ScreenModuleEditorView "IO Field: Single Width; Stacked" 178x111
   IOField "tfLable" at 0,55 size 178x56; FormatPattern ????????????????????????????????????????
      on OnFinishInput: SetBit("Interface.inputFinished")
      Appearance <- "Interface.animate"
      Visibility <- "Interface.visible"
      ProcessValue <- "Interface.value"
      ObjectEnable <- "Interface.enable"
   TextField "iofData" at 0,0 size 178x55; Text 'Text'
      Visibility <- "Interface.visible"
*)

(* ===== HMI "HMI_RT_1" =====
system functions are stored by id; their names below are inferred from use

ScreenModuleEditorView "IO Field: Double Width; Stacked" 370x111
   IOField "tfLable" at 0,55 size 370x56; FormatPattern ????????????????????????????????????????
      on OnFinishInput: SetBit("Interface.inputFinished")
      Appearance <- "Interface.animate"
      ProcessValue <- "Interface.value"
      Visibility <- "Interface.visible"
      ObjectEnable <- "Interface.enable"
   TextField "iofData" at 0,0 size 370x55; Text 'Text'
      Visibility <- "Interface.visible"
*)

(* ===== HMI "HMI_RT_1" =====
system functions are stored by id; their names below are inferred from use

ScreenModuleEditorView "PB: Graphic/Text List" 65x45
   Button "Previous Station Group" at 0,0 size 65x45; TextOff 'Text'
      on Press: function_b14e0dd5("Interface.actuate", 0)
      Visibility <- "Interface.animate"
      ObjectEnable <- "Interface.animate"
      Appearance <- "Interface.animate"
*)

(* ===== HMI "HMI_RT_1" =====
system functions are stored by id; their names below are inferred from use

ScreenModuleEditorView "PB: Graphic/Text List" 65x45
   Button "Previous Station Group" at 0,0 size 65x45; TextOff 'Text'
      on Press: function_b14e0dd5("Interface.actuate", 0)
      Visibility <- "Interface.animate"
      ObjectEnable <- "Interface.animate"
      Appearance <- "Interface.animate"
*)

(* ===== HMI "HMI_RT_1" =====
system functions are stored by id; their names below are inferred from use

ScreenModuleEditorView "PB: Station Comm Status (Text Label)" 180x25
   Button "Station Select" at 0,0 size 180x25; TextOff 'Text'
      on Press: function_b14e0dd5("Interface.actuate", 0)
      Appearance <- "Interface.animate"
      ObjectEnable <- "Interface.enable"
      Visibility <- "Interface.visible"
*)

(* ===== HMI "HMI_RT_1" =====
system functions are stored by id; their names below are inferred from use

ScreenModuleEditorView "PB: Graphic/Text List" 65x45
   Button "Previous Station Group" at 0,0 size 65x45; TextOff 'Text'
      on Press: function_b14e0dd5("Interface.actuate", 0)
      Visibility <- "Interface.animate"
      ObjectEnable <- "Interface.animate"
      Appearance <- "Interface.animate"
*)

(* ===== HMI "HMI_RT_1" =====
system functions are stored by id; their names below are inferred from use

graphic list "Top": 0 '100 x 100 Top'; 1 '100 x 100 Actuated Top'

graphic list "Page Up": 0 '100 x 100 Page Up'; 1 '100 x 100 Actuated Page Up'

graphic list "Line Up": 0 '100 x 100 Line Up'; 1 '100 x 100 Actuated Line Up'

graphic list "Line Down": 0 '100 x 100 Line Down'; 1 '100 x 100 Actuated Line Down'

graphic list "Page Down": 0 '100 x 100 Page Down'; 1 '100 x 100 Actuated Page Down'

graphic list "Bottom": 0 '100 x 100 Bottom'; 1 '100 x 100 Actuated Bottom'

ScreenModuleEditorView "Nav Bar: Horizontal" 600x100
   Button "btnTop" at 1,1 size 98x98; TextOff 'Text'; PictureList "Top"
      on Press: function_b14e0dd5("Interface.top.actuate", 0)
      Visibility <- "Interface.top.visible"
      ObjectEnable <- "Interface.top.enable"
      ProcessValue <- "Interface.top.listSelect"
      Appearance <- "Interface.top.animate"
   Button "btnPageUp" at 101,1 size 98x98; TextOff 'Text'; PictureList "Page Up"
      on Press: function_b14e0dd5("Interface.pageUp.actuate", 0)
      Appearance <- "Interface.pageUp.animate"
      ObjectEnable <- "Interface.pageUp.enable"
      ProcessValue <- "Interface.pageUp.listSelect"
      Visibility <- "Interface.pageUp.visible"
   Button "btnLineUp" at 201,1 size 98x98; TextOff 'Text'; PictureList "Line Up"
      on Press: function_b14e0dd5("Interface.lineUp.actuate", 0)
      Visibility <- "Interface.lineUp.visible"
      ObjectEnable <- "Interface.lineUp.enable"
      ProcessValue <- "Interface.lineUp.listSelect"
      Appearance <- "Interface.lineUp.animate"
   Button "btnLineDown" at 301,1 size 98x98; TextOff 'Text'; PictureList "Line Down"
      on Press: function_b14e0dd5("Interface.lineUp.actuate", 0)
      Appearance <- "Interface.lineDown.animate"
      ObjectEnable <- "Interface.lineDown.enable"
      ProcessValue <- "Interface.lineDown.listSelect"
      Visibility <- "Interface.lineDown.visible"
   Button "btnPageDown" at 401,1 size 98x98; TextOff 'Text'; PictureList "Page Down"
      on Press: function_b14e0dd5("Interface.pageDown.actuate", 0)
      Visibility <- "Interface.pageDown.visible"
      ObjectEnable <- "Interface.pageDown.enable"
      ProcessValue <- "Interface.pageDown.listSelect"
      Appearance <- "Interface.pageDown.animate"
   Button "btnBottom" at 501,1 size 98x98; TextOff 'Text'; PictureList "Bottom"
      on Press: function_b14e0dd5("Interface.pageDown.actuate", 0)
      Appearance <- "Interface.bottom.animate"
      ObjectEnable <- "Interface.bottom.enable"
      ProcessValue <- "Interface.bottom.listSelect"
      Visibility <- "Interface.bottom.visible"
*)

(* ===== HMI "HMI_RT_1" =====
system functions are stored by id; their names below are inferred from use

graphic list "Top": 0 '100 x 100 Top'; 1 '100 x 100 Actuated Top'

graphic list "Page Up": 0 '100 x 100 Page Up'; 1 '100 x 100 Actuated Page Up'

graphic list "Line Up": 0 '100 x 100 Line Up'; 1 '100 x 100 Actuated Line Up'

graphic list "Line Down": 0 '100 x 100 Line Down'; 1 '100 x 100 Actuated Line Down'

graphic list "Page Down": 0 '100 x 100 Page Down'; 1 '100 x 100 Actuated Page Down'

graphic list "Bottom": 0 '100 x 100 Bottom'; 1 '100 x 100 Actuated Bottom'

ScreenModuleEditorView "Nav Bar: Horizontal" 600x100
   Button "btnTop" at 1,1 size 98x98; TextOff 'Text'; PictureList "Top"
      on Press: function_b14e0dd5("Interface.top_actuate", 0)
      Appearance <- "Interface.top_animate"
      ObjectEnable <- "Interface.top_enable"
      Visibility <- "Interface.top_visible"
   Button "btnPageUp" at 101,1 size 98x98; TextOff 'Text'; PictureList "Page Up"
      on Press: function_b14e0dd5("Interface.page_up_actuate", 0)
      Visibility <- "Interface.page_up_visible"
      ObjectEnable <- "Interface.page_up_enable"
      Appearance <- "Interface.page_up_animate"
   Button "btnLineUp" at 201,1 size 98x98; TextOff 'Text'; PictureList "Line Up"
      on Press: function_b14e0dd5("Interface.line_up_actuate", 0)
      Visibility <- "Interface.line_up_visible"
      ObjectEnable <- "Interface.line_up_enable"
      Appearance <- "Interface.line_up_animate"
   Button "btnLineDown" at 301,1 size 98x98; TextOff 'Text'; PictureList "Line Down"
      on Press: function_b14e0dd5("Interface.line_down_actuate", 0)
      Appearance <- "Interface.line_down_animate"
      ObjectEnable <- "Interface.line_down_enable"
      Visibility <- "Interface.line_down_visible"
   Button "btnPageDown" at 401,1 size 98x98; TextOff 'Text'; PictureList "Page Down"
      on Press: function_b14e0dd5("Interface.page_down_actuate", 0)
      Visibility <- "Interface.page_down_visible"
      ObjectEnable <- "Interface.page_down_enable"
      Appearance <- "Interface.page_down_animate"
   Button "btnBottom" at 501,1 size 98x98; TextOff 'Text'; PictureList "Bottom"
      on Press: function_b14e0dd5("Interface.botttom_actuate", 0)
      Appearance <- "Interface.botttom_animate"
      ObjectEnable <- "Interface.botttom_enable"
      Visibility <- "Interface.botttom_visible"
*)

(* ===== HMI "HMI_RT_1" =====
system functions are stored by id; their names below are inferred from use

graphic list "Top": 0 '100 x 100 Top'; 1 '100 x 100 Actuated Top'

graphic list "Page Up": 0 '100 x 100 Page Up'; 1 '100 x 100 Actuated Page Up'

graphic list "Line Up": 0 '100 x 100 Line Up'; 1 '100 x 100 Actuated Line Up'

graphic list "Line Down": 0 '100 x 100 Line Down'; 1 '100 x 100 Actuated Line Down'

graphic list "Page Down": 0 '100 x 100 Page Down'; 1 '100 x 100 Actuated Page Down'

graphic list "Bottom": 0 '100 x 100 Bottom'; 1 '100 x 100 Actuated Bottom'

ScreenModuleEditorView "Nav Bar: Vertical" 100x600
   Button "btnTop" at 1,1 size 98x98; TextOff 'Text'; PictureList "Top"
      on Press: function_b14e0dd5("Interface.top_actuate", 0)
      Appearance <- "Interface.top_animate"
      ObjectEnable <- "Interface.top_enable"
      Visibility <- "Interface.top_visible"
   Button "btnPageUp" at 1,101 size 98x98; TextOff 'Text'; PictureList "Page Up"
      on Press: function_b14e0dd5("Interface.page_up_actuate", 0)
      Visibility <- "Interface.page_up_visible"
      ObjectEnable <- "Interface.page_up_enable"
      Appearance <- "Interface.page_up_animate"
   Button "btnLineUp" at 1,201 size 98x98; TextOff 'Text'; PictureList "Line Up"
      on Press: function_b14e0dd5("Interface.line_up_actuate", 0)
      Appearance <- "Interface.line_up_animate"
      ObjectEnable <- "Interface.line_up_enable"
      Visibility <- "Interface.line_up_visible"
   Button "btnLineDown" at 1,301 size 98x98; TextOff 'Text'; PictureList "Line Down"
      on Press: function_b14e0dd5("Interface.line_down_actuate", 0)
      Visibility <- "Interface.line_down_visible"
      ObjectEnable <- "Interface.line_down_enable"
      Appearance <- "Interface.line_down_animate"
   Button "btnPageDown" at 1,401 size 98x98; TextOff 'Text'; PictureList "Page Down"
      on Press: function_b14e0dd5("Interface.page_down_actuate", 0)
      Appearance <- "Interface.page_down_animate"
      ObjectEnable <- "Interface.page_down_enable"
      Visibility <- "Interface.page_down_visible"
   Button "btnBottom" at 1,501 size 98x98; TextOff 'Text'; PictureList "Bottom"
      on Press: SetBit("Interface.bottom_actuate")
      Visibility <- "Interface.bottom_visible"
      ObjectEnable <- "Interface.bottom_enable"
      Appearance <- "Interface.bottom_animate"
*)

(* ===== HMI "HMI_RT_1" =====
system functions are stored by id; their names below are inferred from use

graphic list "Top": 0 '100 x 100 Top'; 1 '100 x 100 Actuated Top'

graphic list "Page Up": 0 '100 x 100 Page Up'; 1 '100 x 100 Actuated Page Up'

graphic list "Line Up": 0 '100 x 100 Line Up'; 1 '100 x 100 Actuated Line Up'

graphic list "Line Down": 0 '100 x 100 Line Down'; 1 '100 x 100 Actuated Line Down'

graphic list "Page Down": 0 '100 x 100 Page Down'; 1 '100 x 100 Actuated Page Down'

graphic list "Bottom": 0 '100 x 100 Bottom'; 1 '100 x 100 Actuated Bottom'

ScreenModuleEditorView "Nav Bar: Horizontal" 600x100
   Button "btnTop" at 1,1 size 98x98; TextOff 'Text'; PictureList "Top"
      on Press: function_b14e0dd5("Interface.top_actuate", 0)
      Appearance <- "Interface.top_animate"
      ObjectEnable <- "Interface.top_enable"
      Visibility <- "Interface.top_visible"
   Button "btnPageUp" at 101,1 size 98x98; TextOff 'Text'; PictureList "Page Up"
      on Press: function_b14e0dd5("Interface.page_up_actuate", 0)
      Visibility <- "Interface.page_up_visible"
      ObjectEnable <- "Interface.page_up_enable"
      Appearance <- "Interface.page_up_animate"
   Button "btnLineUp" at 201,1 size 98x98; TextOff 'Text'; PictureList "Line Up"
      on Press: function_b14e0dd5("Interface.line_up_actuate", 0)
      Visibility <- "Interface.line_up_visible"
      ObjectEnable <- "Interface.line_up_enable"
      Appearance <- "Interface.line_up_animate"
   Button "btnLineDown" at 301,1 size 98x98; TextOff 'Text'; PictureList "Line Down"
      on Press: function_b14e0dd5("Interface.line_down_actuate", 0)
      Appearance <- "Interface.line_down_animate"
      ObjectEnable <- "Interface.line_down_enable"
      Visibility <- "Interface.line_down_visible"
   Button "btnPageDown" at 401,1 size 98x98; TextOff 'Text'; PictureList "Page Down"
      on Press: function_b14e0dd5("Interface.page_down_actuate", 0)
      Visibility <- "Interface.page_down_visible"
      ObjectEnable <- "Interface.page_down_enable"
      Appearance <- "Interface.page_down_animate"
   Button "btnBottom" at 501,1 size 98x98; TextOff 'Text'; PictureList "Bottom"
      on Press: function_b14e0dd5("Interface.bottom_actuate", 0)
      Visibility <- "Interface.bottom_visible"
      ObjectEnable <- "Interface.bottom_enable"
      Appearance <- "Interface.bottom_animate"
*)

(* ===== HMI "HMI_RT_1" =====
system functions are stored by id; their names below are inferred from use

graphic list "Top": 0 '100 x 100 Top'; 1 '100 x 100 Actuated Top'

graphic list "Page Up": 0 '100 x 100 Page Up'; 1 '100 x 100 Actuated Page Up'

graphic list "Line Up": 0 '100 x 100 Line Up'; 1 '100 x 100 Actuated Line Up'

graphic list "Line Down": 0 '100 x 100 Line Down'; 1 '100 x 100 Actuated Line Down'

graphic list "Page Down": 0 '100 x 100 Page Down'; 1 '100 x 100 Actuated Page Down'

graphic list "Bottom": 0 '100 x 100 Bottom'; 1 '100 x 100 Actuated Bottom'

ScreenModuleEditorView "Nav Bar: Horizontal" 600x100
   Button "btnTop" at 1,1 size 98x98; TextOff 'Text'; PictureList "Top"
      on Press: function_b14e0dd5("Interface.top_actuate", 0)
      Appearance <- "Interface.top_animate"
      ObjectEnable <- "Interface.top_enable"
      Visibility <- "Interface.top_visible"
      ProcessValue <- "Interface.top_list_select"
   Button "btnPageUp" at 101,1 size 98x98; TextOff 'Text'; PictureList "Page Up"
      on Press: function_b14e0dd5("Interface.page_up_actuate", 0)
      Visibility <- "Interface.page_up_visible"
      ObjectEnable <- "Interface.page_up_enable"
      Appearance <- "Interface.page_up_animate"
      ProcessValue <- "Interface.page_up_list_select"
   Button "btnLineUp" at 201,1 size 98x98; TextOff 'Text'; PictureList "Line Up"
      on Press: function_b14e0dd5("Interface.line_up_actuate", 0)
      Visibility <- "Interface.line_up_visible"
      ObjectEnable <- "Interface.line_up_enable"
      Appearance <- "Interface.line_up_animate"
      ProcessValue <- "Interface.line_up_list_select"
   Button "btnLineDown" at 301,1 size 98x98; TextOff 'Text'; PictureList "Line Down"
      on Press: function_b14e0dd5("Interface.line_down_actuate", 0)
      Appearance <- "Interface.line_down_animate"
      ObjectEnable <- "Interface.line_down_enable"
      Visibility <- "Interface.line_down_visible"
      ProcessValue <- "Interface.line_down_list_select"
   Button "btnPageDown" at 401,1 size 98x98; TextOff 'Text'; PictureList "Page Down"
      on Press: function_b14e0dd5("Interface.page_down_actuate", 0)
      Visibility <- "Interface.page_down_visible"
      ObjectEnable <- "Interface.page_down_enable"
      Appearance <- "Interface.page_down_animate"
      ProcessValue <- "Interface.page_down_list_select"
   Button "btnBottom" at 501,1 size 98x98; TextOff 'Text'; PictureList "Bottom"
      on Press: function_b14e0dd5("Interface.bottom_actuate", 0)
      Visibility <- "Interface.bottom_visible"
      ObjectEnable <- "Interface.bottom_enable"
      Appearance <- "Interface.bottom_animate"
      ProcessValue <- "Interface.bottom_list_select"
*)

(* ===== HMI "HMI_RT_1" =====
system functions are stored by id; their names below are inferred from use

ScreenModuleEditorView "PB: Dynamic Text Label" 100x100
   Button "pbActuate" at 0,0 size 100x100; TextOff 'Text'
      on Release: ResetBit("Interface.actuate")
      on Press: SetBit("Interface.actuate")
      Visibility <- "Interface.visible"
      ObjectEnable <- "Interface.enable"
   TextField "tfDisplay" at 0,0 size 100x100; Text 'Text'
      Visibility <- "Interface.visible"
      Appearance <- "Interface.animate"
*)

(* ===== HMI "HMI_RT_1" =====
system functions are stored by id; their names below are inferred from use

ScreenModuleEditorView "PB: Dynamic Text Label" 100x100
   Button "pbActuate" at 0,0 size 100x100; TextOff 'Text'
      on Release: ResetBit("Interface.actuate")
      on Press: SetBit("Interface.actuate")
      Visibility <- "Interface.visible"
      ObjectEnable <- "Interface.enable"
   TextField "tfDisplay" at 0,0 size 100x100; Text 'Text'
      Visibility <- "Interface.visible"
      Appearance <- "Interface.animate"
*)

(* ===== HMI "HMI_RT_1" =====
system functions are stored by id; their names below are inferred from use

ScreenModuleEditorView "PB: Static Text Label" 274x45
   Button "Select All Stations" at 0,0 size 274x45; TextOff 'Text'
      on Press: function_b14e0dd5("Interface.actuate", 0)
      Appearance <- "Interface.animate"
      ObjectEnable <- "Interface.enable"
      Visibility <- "Interface.visible"
*)

(* ===== HMI "HMI_RT_1" =====
system functions are stored by id; their names below are inferred from use

ScreenModuleEditorView "PB: Dynamic Text Label" 100x100
   Button "pbActuate" at 0,0 size 100x100; TextOff 'Text'
      on Release: ResetBit("Interface.actuate")
      on Press: SetBit("Interface.actuate")
      Visibility <- "Interface.visible"
      ObjectEnable <- "Interface.enable"
   TextField "tfDisplay" at 0,0 size 100x100; Text 'Text'
      Visibility <- "Interface.visible"
      Appearance <- "Interface.animate"
*)

(* ===== HMI "HMI_RT_1" =====
system functions are stored by id; their names below are inferred from use

ScreenModuleEditorView "PB: Dynamic Text Label" 100x100
   Button "pbActuate" at 0,0 size 100x100; TextOff 'Text'
      on Release: ResetBit("Interface.actuate")
      on Press: SetBit("Interface.actuate")
      Visibility <- "Interface.visible"
      ObjectEnable <- "Interface.enable"
   TextField "tfDisplay" at 0,0 size 100x100; Text 'Text'
      Visibility <- "Interface.visible"
      Appearance <- "Interface.animate"
*)

(* ===== HMI "HMI_RT_1" =====
system functions are stored by id; their names below are inferred from use

ScreenModuleEditorView "PB: Dynamic Text Label" 100x100
   Button "pbActuate" at 0,0 size 100x100; TextOff 'Text'
      on Release: ResetBit("Interface.actuate")
      on Press: SetBit("Interface.actuate")
      Visibility <- "Interface.visible"
      ObjectEnable <- "Interface.enable"
   TextField "tfDisplay" at 0,0 size 100x100; Text 'Text'
      Visibility <- "Interface.visible"
      Appearance <- "Interface.animate"
*)

(* ===== HMI "HMI_RT_1" =====
system functions are stored by id; their names below are inferred from use

ScreenModuleEditorView "PB: Dynamic Text Label" 100x100
   Button "pbActuate" at 0,0 size 100x100; TextOff 'Text'
      on Release: ResetBit("Interface.actuate")
      on Press: SetBit("Interface.actuate")
      Visibility <- "Interface.visible"
      ObjectEnable <- "Interface.enable"
   TextField "tfDisplay" at 0,0 size 100x100; Text 'Text'
      Visibility <- "Interface.visible"
      Appearance <- "Interface.animate"
*)

(* ===== HMI "HMI_RT_1" =====
system functions are stored by id; their names below are inferred from use

ScreenModuleEditorView "PB: Static Text Label" 274x45
   Button "Select All Stations" at 0,0 size 274x45; TextOff 'Text'
      on Press: function_b14e0dd5("Interface.actuate", 0)
      Appearance <- "Interface.animate"
      ObjectEnable <- "Interface.enable"
      Visibility <- "Interface.visible"
*)

(* ===== HMI "HMI_RT_1" =====
system functions are stored by id; their names below are inferred from use

graphic list "Top": 0 '100 x 100 Top'; 1 '100 x 100 Actuated Top'

graphic list "Page Up": 0 '100 x 100 Page Up'; 1 '100 x 100 Actuated Page Up'

graphic list "Line Up": 0 '100 x 100 Line Up'; 1 '100 x 100 Actuated Line Up'

graphic list "Line Down": 0 '100 x 100 Line Down'; 1 '100 x 100 Actuated Line Down'

graphic list "Page Down": 0 '100 x 100 Page Down'; 1 '100 x 100 Actuated Page Down'

graphic list "Bottom": 0 '100 x 100 Bottom'; 1 '100 x 100 Actuated Bottom'

ScreenModuleEditorView "Nav Bar: Vertical" 100x600
   Button "btnTop" at 1,1 size 98x98; TextOff 'Text'; PictureList "Top"
      on Press: function_b14e0dd5("Interface.top_actuate", 0)
      Appearance <- "Interface.top_animate"
      ObjectEnable <- "Interface.top_enable"
      Visibility <- "Interface.top_visible"
      ProcessValue <- "Interface.top_list_select"
   Button "btnPageUp" at 1,101 size 98x98; TextOff 'Text'; PictureList "Page Up"
      on Press: function_b14e0dd5("Interface.page_up_actuate", 0)
      Visibility <- "Interface.page_up_visible"
      ObjectEnable <- "Interface.page_up_enable"
      Appearance <- "Interface.page_up_animate"
      ProcessValue <- "Interface.page_up_list_select"
   Button "btnLineUp" at 1,201 size 98x98; TextOff 'Text'; PictureList "Line Up"
      on Press: function_b14e0dd5("Interface.line_up_actuate", 0)
      Appearance <- "Interface.line_up_animate"
      ObjectEnable <- "Interface.line_up_enable"
      Visibility <- "Interface.line_up_visible"
      ProcessValue <- "Interface.line_up_list_select"
   Button "btnLineDown" at 1,301 size 98x98; TextOff 'Text'; PictureList "Line Down"
      on Press: function_b14e0dd5("Interface.line_down_actuate", 0)
      Visibility <- "Interface.line_down_visible"
      ObjectEnable <- "Interface.line_down_enable"
      Appearance <- "Interface.line_down_animate"
      ProcessValue <- "Interface.line_down_list_select"
   Button "btnPageDown" at 1,401 size 98x98; TextOff 'Text'; PictureList "Page Down"
      on Press: function_b14e0dd5("Interface.page_down_actuate", 0)
      Appearance <- "Interface.page_down_animate"
      ObjectEnable <- "Interface.page_down_enable"
      Visibility <- "Interface.page_down_visible"
      ProcessValue <- "Interface.page_down_list_select"
   Button "btnBottom" at 1,501 size 98x98; TextOff 'Text'; PictureList "Bottom"
      on Press: SetBit("Interface.bottom_actuate")
      Visibility <- "Interface.bottom_visible"
      ObjectEnable <- "Interface.bottom_enable"
      Appearance <- "Interface.bottom_animate"
      ProcessValue <- "Interface.bottom_list_select"
*)

(* ===== HMI "HMI_RT_1" =====
system functions are stored by id; their names below are inferred from use

graphic list "Top": 0 '100 x 100 Top'; 1 '100 x 100 Actuated Top'

graphic list "Page Up": 0 '100 x 100 Page Up'; 1 '100 x 100 Actuated Page Up'

graphic list "Line Up": 0 '100 x 100 Line Up'; 1 '100 x 100 Actuated Line Up'

graphic list "Line Down": 0 '100 x 100 Line Down'; 1 '100 x 100 Actuated Line Down'

graphic list "Page Down": 0 '100 x 100 Page Down'; 1 '100 x 100 Actuated Page Down'

graphic list "Bottom": 0 '100 x 100 Bottom'; 1 '100 x 100 Actuated Bottom'

ScreenModuleEditorView "Nav Bar: Vertical" 100x600
   Button "btnTop" at 1,1 size 98x98; TextOff 'Text'; PictureList "Top"
      on Press: function_b14e0dd5("Interface.top_actuate", 0)
      Appearance <- "Interface.top_animate"
      ObjectEnable <- "Interface.top_enable"
      ProcessValue <- "Interface.top_list_select"
      Visibility <- "Interface.top_visible"
   Button "btnPageUp" at 1,101 size 98x98; TextOff 'Text'; PictureList "Page Up"
      on Press: function_b14e0dd5("Interface.page_up_actuate", 0)
      Visibility <- "Interface.page_up_visible"
      ObjectEnable <- "Interface.page_up_enable"
      ProcessValue <- "Interface.page_up_list_select"
      Appearance <- "Interface.page_up_animate"
   Button "btnLineUp" at 1,201 size 98x98; TextOff 'Text'; PictureList "Line Up"
      on Press: function_b14e0dd5("Interface.line_up_actuate", 0)
      Appearance <- "Interface.line_up_animate"
      ObjectEnable <- "Interface.line_up_enable"
      ProcessValue <- "Interface.line_up_list_select"
      Visibility <- "Interface.line_up_visible"
   Button "btnLineDown" at 1,301 size 98x98; TextOff 'Text'; PictureList "Line Down"
      on Press: function_b14e0dd5("Interface.line_down_actuate", 0)
      Visibility <- "Interface.line_down_visible"
      ObjectEnable <- "Interface.line_down_enable"
      ProcessValue <- "Interface.line_down_list_select"
      Appearance <- "Interface.line_down_animate"
   Button "btnPageDown" at 1,401 size 98x98; TextOff 'Text'; PictureList "Page Down"
      on Press: function_b14e0dd5("Interface.page_down_actuate", 0)
      Appearance <- "Interface.page_down_animate"
      ObjectEnable <- "Interface.page_down_enable"
      ProcessValue <- "Interface.page_down_list_select"
      Visibility <- "Interface.page_down_visible"
   Button "btnBottom" at 1,501 size 98x98; TextOff 'Text'; PictureList "Bottom"
      on Press: function_b14e0dd5("Interface.bottom_actuate", 0)
      Visibility <- "Interface.bottom_visible"
      ObjectEnable <- "Interface.bottom_enable"
      ProcessValue <- "Interface.bottom_list_select"
      Appearance <- "Interface.bottom_animate"
*)

(* ===== HMI "HMI_RT_1" =====
system functions are stored by id; their names below are inferred from use

ScreenModuleEditorView "IO Field: Single Width; Stacked" 178x111
   IOField "tfLable" at 0,55 size 178x56; FormatPattern ????????????????????????????????????????
      on OnFinishInput: SetBit("Interface.input_finished")
      Appearance <- "Interface.animate"
      Visibility <- "Interface.visible"
      ObjectEnable <- "Interface.enable"
      ProcessValue <- "Interface.value"
   TextField "iofData" at 0,0 size 178x55; Text 'Text'
      Visibility <- "Interface.visible"
      Appearance <- "Interface.animate"
*)

(* ===== HMI "HMI_RT_1" =====
system functions are stored by id; their names below are inferred from use

ScreenModuleEditorView "IO Field: Single Width; Stacked" 178x111
   IOField "tfLable" at 0,55 size 178x56; FormatPattern ????????????????????????????????????????
      on OnFinishInput: SetBit("Interface.input_finished")
      Appearance <- "Interface.animate"
      Visibility <- "Interface.visible"
      ProcessValue <- "Interface.value"
      ObjectEnable <- "Interface.enable"
   TextField "iofData" at 0,0 size 178x55; Text 'Text'
      Visibility <- "Interface.visible"
      Appearance <- "Interface.animate"
*)

(* ===== HMI "HMI_RT_1" =====
system functions are stored by id; their names below are inferred from use

ScreenModuleEditorView "IO Field: Single Width; Stacked" 178x111
   IOField "tfLable" at 0,55 size 178x56; FormatPattern ????????????????????????????????????????
      on OnFinishInput: SetBit("Interface.input_finished")
      Appearance <- "Interface.animate"
      Visibility <- "Interface.visible"
      ObjectEnable <- "Interface.enable"
      ProcessValue <- "Interface.value"
   TextField "iofData" at 0,0 size 178x55; Text 'Text'
      Visibility <- "Interface.visible"
      Appearance <- "Interface.animate"
*)

(* ===== HMI "HMI_RT_1" =====
system functions are stored by id; their names below are inferred from use

ScreenModuleEditorView "IO Field: Single Width; Stacked" 178x111
   IOField "tfLable" at 0,55 size 178x56; FormatPattern ????????????????????????????????????????
      on OnFinishInput: SetBit("Interface.input_finished")
      Appearance <- "Interface.animate"
      Visibility <- "Interface.visible"
      ProcessValue <- "Interface.value"
      ObjectEnable <- "Interface.enable"
   TextField "iofData" at 0,0 size 178x55; Text 'Text'
      Visibility <- "Interface.visible"
      Appearance <- "Interface.animate"
*)

(* ===== HMI "HMI_RT_1" =====
system functions are stored by id; their names below are inferred from use

ScreenModuleEditorView "IO Field: Double Width; Stacked" 370x111
   IOField "tfLable" at 0,55 size 370x56; FormatPattern ????????????????????????????????????????
      on OnFinishInput: SetBit("Interface.inputFinished")
      Appearance <- "Interface.animate"
      ProcessValue <- "Interface.value"
      ObjectEnable <- "Interface.enable"
      Visibility <- "Interface.visible"
   TextField "iofData" at 0,0 size 370x55; Text 'Text'
      Visibility <- "Interface.visible"
      Appearance <- "Interface.animate"
*)

(* ===== HMI "HMI_RT_1" =====
system functions are stored by id; their names below are inferred from use

ScreenModuleEditorView "IO Field: Single Width; Stacked" 178x111
   IOField "tfLable" at 0,55 size 178x56; FormatPattern ????????????????????????????????????????
      on OnFinishInput: SetBit("Interface.input_finished")
      Appearance <- "Interface.animate"
      Visibility <- "Interface.visible"
      ObjectEnable <- "Interface.enable"
      ProcessValue <- "Interface.value"
   TextField "iofData" at 0,0 size 178x55; Text 'Text'
      Visibility <- "Interface.visible"
      Appearance <- "Interface.animate"
*)

(* ===== HMI "HMI_RT_1" =====
system functions are stored by id; their names below are inferred from use

ScreenModuleEditorView "IO Field: Single Width; Stacked" 178x111
   IOField "tfLable" at 0,55 size 178x56; FormatPattern ????????????????????????????????????????
      on OnFinishInput: SetBit("Interface.input_finished")
      Appearance <- "Interface.animate"
      Visibility <- "Interface.visible"
      ProcessValue <- "Interface.value"
      ObjectEnable <- "Interface.enable"
   TextField "iofData" at 0,0 size 178x55; Text 'Text'
      Visibility <- "Interface.visible"
      Appearance <- "Interface.animate"
*)

(* ===== HMI "HMI_RT_1" =====
system functions are stored by id; their names below are inferred from use

ScreenModuleEditorView "IO Field: Double Width; Stacked" 370x111
   IOField "tfLable" at 0,55 size 370x56; FormatPattern ????????????????????????????????????????
      on OnFinishInput: SetBit("Interface.inputFinished")
      Appearance <- "Interface.animate"
      Visibility <- "Interface.visible"
      ProcessValue <- "Interface.value"
      ObjectEnable <- "Interface.enable"
   TextField "iofData" at 0,0 size 370x55; Text 'Text'
      Visibility <- "Interface.visible"
      Appearance <- "Interface.animate"
*)